         reasonOutputSwitchedOff2 : Int;   // 0=output current>limit and output current<1,5xlimit for more than 5sec; 1=current output>1,5xlimit; 2=total overload; 3=Uin<19,4V and output current>limit; 4=Uin<15V; 5=Uin>30V; 6=device overtemperature; 8 to 14=Reserve; 15=default (no automatically switched off)
         reasonOutputSwitchedOff3 : Int;   // 0=output current>limit and output current<1,5xlimit for more than 5sec; 1=current output>1,5xlimit; 2=total overload; 3=Uin<19,4V and output current>limit; 4=Uin<15V; 5=Uin>30V; 6=device overtemperature; 8 to 14=Reserve; 15=default (no automatically switched off)
         reasonOutputSwitchedOff4 : Int;   // 0=output current>limit and output current<1,5xlimit for more than 5sec; 1=current output>1,5xlimit; 2=total overload; 3=Uin<19,4V and output current>limit; 4=Uin<15V; 5=Uin>30V; 6=device overtemperature; 8 to 14=Reserve; 15=default (no automatically switched off)
         reasonOutputSwitchedOff5 : Int;   // 0=output current>limit and output current<1,5xlimit for more than 5sec; 1=current output>1,5xlimit; 2=total overload; 3=Uin<19,4V and output current>limit; 4=Uin<15V; 5=Uin>30V; 6=device overtemperature; 8 to 14=Reserve; 15=default (no automatically switched off)
         reasonOutputSwitchedOff6 : Int;   // 0=output current>limit and output current<1,5xlimit for more than 5sec; 1=current output>1,5xlimit; 2=total overload; 3=Uin<19,4V and output current>limit; 4=Uin<15V; 5=Uin>30V; 6=device overtemperature; 8 to 14=Reserve; 15=default (no automatically switched off)
         reasonOutputSwitchedOff7 : Int;   // 0=output current>limit and output current<1,5xlimit for more than 5sec; 1=current output>1,5xlimit; 2=total overload; 3=Uin<19,4V and output current>limit; 4=Uin<15V; 5=Uin>30V; 6=device overtemperature; 8 to 14=Reserve; 15=default (no automatically switched off)
         reasonOutputSwitchedOff8 : Int;   // 0=output current>limit and output current<1,5xlimit for more than 5sec; 1=current output>1,5xlimit; 2=total overload; 3=Uin<19,4V and output current>limit; 4=Uin<15V; 5=Uin>30V; 6=device overtemperature; 8 to 14=Reserve; 15=default (no automatically switched off)
         nominalOutputCurrent : Int;   // nominal output current
         outputNumber : Int;   // number of outputs (4 or 8)
         productState : Int;   // product state
         firmwareVersion : Int;   // frimware version
         startup : Int;   // 0=load dependent startup; 1=startup time tag 25ms; 2=startup time tag 200ms; 3=startup time tag 500ms
         setReset : Bool;
         stateReset : Bool;
         stateNoCommunication : Bool;
         articleNumber : String;   // article number
         serialNumber : String;   // serial number
      END_STRUCT;
      statIndexResetBitArray : Int;
      statInit : Bool;
      statArticleNumber : Array[1..18] of Char;
      statArticleNumberOld : Array[1..18] of Char;
      statSerialNumber : Array[1..13] of Char;
      statSerialNumberOld : Array[1..13] of Char;
      statVarianten11String : String[2];
      statInnovationenString : String[2];
      statArticleNumberChanged : Bool;
      statErrorFrameContent : Bool;
      statErrorFrameID : Bool;
      statErrorFrameLength : Bool;
      statErrorDevice : Bool;
      statIndexArticleNumber : Int := 1;
      statIndexSerialNumber : Int := 1;
      statNewArticleNumberDetected : Bool;
      statNewSerialNumberDetected : Bool;
      instTimerReset : TON_TIME;
      statCntReason : Int;
      statCntCurrentLimit : Int;
   END_VAR
   VAR_TEMP
      tempLatchTime : Time;
      tempRetval : Word;
      tempRetvalSysTime : Int;
      tempRetvalSysPosEdge : Int;
      tempRetvalSysNegEdge : Int;
   END_VAR
   VAR CONSTANT
      CONST_POS_EDGE : Int := 15;
      CONST_NEG_EDGE : Int := 16;
      STATE_IDLE : Int := 1;
      STATE_EVALUATION : Int := 2;
      STATE_ERROR : Int := 3;
      CONST_DWORD_0 : DWord := 16#0000_0000;
      CONST_WORD_0 : Word := 16#0000;
      CONST_BYTE_0 : Byte := 16#00;
      CONST_INT_0 : Int := 0;
      CONST_INT_1 : Int := 1;
      CONST_TIME_0 : Time := T#0MS;
      CONST_TIME_WAIT : Time := T#65MS;
      CONST_SYS_TIMER : Time := T#4S;
      CONST_WATCHDOG_TIMER : Time := T#9S;
      CONST_INIT_TIMER : Time := T#4S;
      CONST_RESET_TIMER : Time := T#50ms;
      CONST_START_IMPULSE_MIN : Time := T#126MS;
      CONST_START_IMPULSE_MAX : Time := T#175MS;
      CONST_IMPULSE_MIN : Time := T#25MS;
      CONST_IMPULSE_MAX : Time := T#125MS;
      CONST_PAUSE_MAX : Time := T#125MS;
      CONST_PAUSE_MIN : Time := T#25MS;
      CONST_START_CNT_INDEX0 : Int := 0;
      CONST_START_CNT_INDEX1 : Int := 1;
      CONST_END_CNT_INDEX63 : Int := 63;
      CONST_END_CNT_INDEX31 : Int := 31;
      CONST_END_CNT_INDEX18 : Int := 18;
      CONST_END_CNT_INDEX13 : Int := 13;
      CONST_FRAME_MAX : Time := T#3S_625MS;
      CONST_FRAME_MIN : Time := T#3S_275MS;
      CONST_CNT_BITS_MAX : Int := 32;
      CONST_CNT_PAUSE_MAX : Int := 33;
      CONST_TIME_CYCLE_MAX : Time := T#12MS;
      CONST_ERR_ARTICLE_NUMBER : Word := 16#8007;
      CONST_ERR_FRAME_ID : Word := 16#8006;
      CONST_ERR_DEVICE : Word := 16#8005;
      CONST_ERR_FRAMELENGTH : Word := 16#8004;
      CONST_ERR_FRAMECONTENT : Word := 16#8003;
      CONST_ERR_CYCLE_TIME : Word := 16#8002;
      CONST_ERR_WATCHDOG : Word := 16#8001;
      CONST_CONVERT_CURRENT : Int := 10;
      CONST_NOMINAL_VALUE_DETECT0 : Byte := 16#00;
      CONST_NOMINAL_VALUE_DETECT1 : Byte := 16#01;
      CONST_NOMINAL_VALUE_DETECT2 : Byte := 16#02;
      CONST_NOMINAL_CURRENT3 : Int := 3;
      CONST_NOMINAL_CURRENT5 : Int := 5;
      CONST_NOMINAL_CURRENT10 : Int := 10;
      CONST_NOMINAL_VOLTAGE : Int := 24;
      CONST_YEAR_2019 : Int := 2019;
      CONST_YEAR_2020 : Int := 2020;
      CONST_YEAR_2021 : Int := 2021;
      CONST_YEAR_2022 : Int := 2022;
      CONST_YEAR_2023 : Int := 2023;
      CONST_YEAR_2024 : Int := 2024;
      CONST_YEAR_2025 : Int := 2025;
      CONST_YEAR_2026 : Int := 2026;
      CONST_YEAR_2027 : Int := 2027;
      CONST_YEAR_2028 : Int := 2028;
      CONST_YEAR_2029 : Int := 2029;
      CONST_YEAR_2030 : Int := 2030;
      CONST_YEAR_2031 : Int := 2031;
      CONST_YEAR_2032 : Int := 2032;
      CONST_YEAR_2033 : Int := 2033;
      CONST_YEAR_2034 : Int := 2034;
      CONST_FRAME_ID0 : Int := 0;
      CONST_FRAME_ID1 : Int := 1;
      CONST_FRAME_ID2 : Int := 2;
      CONST_FRAME_ID3 : Int := 3;
      CONST_DEVICE_SEL1200 : Int := 1;
      CONST_DEVICE_SEL1400 : Int := 2;
      CONST_JANUARY : Int := 1;
      CONST_FEBRUARY : Int := 2;
      CONST_MARCH : Int := 3;
      CONST_APRIL : Int := 4;
      CONST_MAY : Int := 5;
      CONST_JUNE : Int := 6;
      CONST_JULY : Int := 7;
      CONST_AUGUST : Int := 8;
      CONST_SEPTEMBER : Int := 9;
      CONST_OCTOBER : Int := 10;
      CONST_NOVEMBER : Int := 11;
      CONST_DECEMBER : Int := 12;
      CONST_ONE_CHANNEL : Int := 0;
      CONST_TWO_CHANNEL : Int := 1;
      CONST_FOUR_CHANNEL : Int := 2;
      CONST_EIGHT_CHANNEL : Int := 3;
      CONST_NO_DESCRIPTION : Int := 4;
      CONST_GLITCH_MAX : Int := 32000;
      CONST_MEASUREMENT_CURRENT : Int := 0;
      CONST_MEASUREMENT_CURRENT_LIMIT : Int := 2;
      CONST_OUTPUT_NUMBER_4 : Int := 4;
      CONST_OUTPUT_NUMBER_8 : Int := 8;
      CONST_POWER_0 : Int := 0;
      CONST_POWER_20 : Int := 20;
      CONST_POWER_50 : Int := 50;
      CONST_POWER_100 : Int := 100;
      CONST_POWER_150 : Int := 150;
      CONST_POWER_250 : Int := 250;
      CONST_POWER_400 : Int := 400;
      CONST_POWER_600 : Int := 600;
      CONST_POWER_1000 : Int := 100;
      CONST_REASON_DEFAULT : Int := 0;
      CONST_STATE_OUT_AUTO_SWITCHED_OFF : Int := 0;
      CONST_STATE_OUT_RESET_POSSIBLE : Int := 1;
      CONST_DEVICE_NAME_DEFAULT : String := 'SEL1200';
      CONST_ARTICLE_NUMBER_DEFAULT : String := '6EP4437-7FB00-0CX0';
      CONST_SERIAL_NUMBER_DEFAULT : String := 'Q6/L1';
      CONST_STATE_OUT_DEFAULT : Int := 0;
      CONST_CURRENT_OUT_DEFAULT : Int := 0;
      CONST_REASON_SWITCHED_OFF_DEFAULT : Int := 0;
      CONST_FW_PRODUCT_STATE_DEFAULT : Int := 1;
      CONST_STARTUP_DEFAULT : Int := 0;
   END_VAR
BEGIN

REGION Network 1 (SCL)
   //=============================================================================
   //SIEMENES AG
   //(c)Copyright 2019 All Rights Reserved
   //-----------------------------------------------------------------------------
   //Library:       LPSU6200_V15.0-0_V1-0-0
   //Tested with:   (S7-1500)
   //Engineering:    TIA Portal V15
   //Restrictions:   call in cyclic interrupt OB with max. 10ms
   //Requirements:
   //Functionality: evaluates the signal of diagnostic interface of SITOP PSU6200 
   //               ....
   //
   //-----------------------------------------------------------------------------
   //Change log table:
   //Version  Date       Expert in charge Changes applied
   //01.00.00 17.01.2019 (DF CS SD CSS KMT KD) First released version
   //=============================================================================


   // Calculate cycle time
   #tempRetvalSysTime := RD_SYS_T(#statTimeSave.sysTime);

   IF #statTimeSave.sysTime > #statTimeSave.sysTimeOld
   THEN
       //Calculate cycle time
       #statTimeSave.deltaSysTime := T_DIFF(IN1 := #statTimeSave.sysTime,
                                            IN2 := #statTimeSave.sysTimeOld);
       #statStartTimerSys := false;
   ELSE
       #statStartTimerSys := true;
       #statTimeSave.sysTimeOld := #statTimeSave.sysTime;
       RETURN;
   END_IF;

   //check cycle time

   IF (#statTimeSave.deltaSysTime >= #CONST_TIME_CYCLE_MAX)
   THEN
       #statCycleTimeNotOk := true;
       #statStartTimerSys := true;
   ELSE
       #statCycleTimeNotOk := false;
       #statStartTimerSys := false;
   END_IF;


   //pos edge detection

   IF #impulse = TRUE
       AND #statImpulseOld = FALSE
   THEN
       #tempRetvalSysPosEdge := RD_SYS_T(#statTimeSave.posEdge);
       #statPosEdgeDetected := true;
       #statPosEdgeDetectedTrigger := true;
       #statEdgeCtrl := #CONST_POS_EDGE;
       #statStartWatchDogTimerPos := true;
       #statStartWatchDogTimerNeg := false;
       #HMI.stateNoCommunication := false;

       IF #statBusy = FALSE
       THEN
           #statInit := false;
           #statBusy := true;
           #statDone := false;
           #statError := false;
           #statStatus := #CONST_WORD_0;
       END_IF;

       IF #statCycleTimeNotOk = FALSE
       THEN
           #statStateIndex := #STATE_EVALUATION;
       END_IF;

   END_IF;

   //neg edge detection

   IF #impulse = false
       AND #statImpulseOld = true
   THEN
       #tempRetvalSysNegEdge := RD_SYS_T(#statTimeSave.negEdge);
       #statNegEdgeDetected := true;
       #statNegEdgeDetectedTrigger := true;
       #statEdgeCtrl := #CONST_NEG_EDGE;
       #statStartWatchDogTimerNeg := true;
       #statStartWatchDogTimerPos := false;

       IF #statCycleTimeNotOk = FALSE
       THEN
           #statStateIndex := #STATE_EVALUATION;
       END_IF;

   END_IF;

   IF #statPosEdgeDetected = FALSE
       AND #statNegEdgeDetected = FALSE
   THEN
       #statStartWatchDogTimerPos := true;
       #statStartWatchDogTimerNeg := true;
   END_IF;


   CASE #statStateIndex OF
       #STATE_IDLE:  // State IDLE

           #statError := false;
           #statErrorInt := false;
           #statDone := false;
           #statBusy := false;
           #statStatus := #CONST_WORD_0;
           #statFrame := #CONST_DWORD_0;
           #statInit := false;
           #error := false;
           #done := false;
           #busy := false;
           #status := #CONST_WORD_0;
           #frame := #CONST_DWORD_0;

           #statNoEvaluation := false;
           #statFrameEvaluationStopp := false;
           #statStartTimerWait := false;
           #statCycleTimeNotOk := false;
           #statPosEdgeDetected := false;
           #statNegEdgeDetected := false;
           #HMI.stateNoCommunication := false;

           FOR #statIndexResetBitArray := #CONST_START_CNT_INDEX0 TO #CONST_END_CNT_INDEX31 DO
               // Statement section FOR
               #statArrayBits[#statIndexResetBitArray] := false;
           END_FOR;


       #STATE_EVALUATION:

           IF #statPosEdgeDetected = TRUE
               AND #statNegEdgeDetected = true
           THEN


               // Delta Time calculation

               IF #statEdgeCtrl = #CONST_POS_EDGE
               THEN
                   #statPauseDetected := true;

                   // time of pause
                   #statTimeSave.deltaTimePause := T_DIFF(IN1 := #statTimeSave.posEdge,
                                                          IN2 := #statTimeSave.negEdge);

                   //check time of pause
                   IF #statTimeSave.deltaTimePause < #CONST_TIME_0
                   THEN
                       #statErrorFrameContent := TRUE;
                   ELSIF (#statTimeSave.deltaTimePause < #CONST_PAUSE_MIN)
                       OR (#statTimeSave.deltaTimePause > #CONST_PAUSE_MAX)
                   THEN
                       #statErrorFrameContent := TRUE;
                   END_IF;

                   #statNegEdgeDetected := false;
               END_IF;

               IF #statEdgeCtrl = #CONST_NEG_EDGE
               THEN
                   #statImpulseDetected := true;

                   // time of impulse
                   #statTimeSave.deltaTimeImpulse := T_DIFF(IN1 := #statTimeSave.negEdge,
                                                            IN2 := #statTimeSave.posEdge);

                   //check time of impulse

                   IF #statTimeSave.deltaTimeImpulse < #CONST_TIME_0
                   THEN
                       #statErrorFrameContent := TRUE;

                   ELSIF (#statTimeSave.deltaTimeImpulse < #CONST_IMPULSE_MIN)
                       OR (#statTimeSave.deltaTimeImpulse > #CONST_START_IMPULSE_MAX)
                   THEN
                       #statErrorFrameContent := TRUE;
                   END_IF;

                   #statPosEdgeDetected := false;
               END_IF;

           END_IF;

           //Startbit detection
           IF (#statTimeSave.deltaTimeImpulse >= #CONST_START_IMPULSE_MIN)
               AND (#statTimeSave.deltaTimeImpulse <= #CONST_START_IMPULSE_MAX)
               AND (#statImpulseDetected = true)
           THEN
               #statImpulseDetected := false;
               #statIndexImpulse := #CONST_INT_1;
               #statIndexPause := #CONST_INT_0;
               #statFrameEvaluationStopp := false;
               #statCntBits := #CONST_INT_0;
               #statCntImpulse := #CONST_INT_0;
               #statCntPause := #CONST_INT_0;
               #statTimeSave.timeIpulse := #CONST_TIME_0;
               #statTimeSave.timePause := #CONST_TIME_0;
               #statIndexAddTime := #CONST_INT_0;

               //check frame length
               FOR #statIndexAddTime := #CONST_START_CNT_INDEX0 TO #CONST_END_CNT_INDEX63 BY 1 DO
                   #statTimeSave.timeIpulse := #statTimeSave.timeIpulse + #statArrayImpulse[#statIndexAddTime];
                   #statTimeSave.timePause := #statTimeSave.timePause + #statArrayPause[#statIndexAddTime];
               END_FOR;

               #statTimeSave.timeFrame := #statTimeSave.timeIpulse + #statTimeSave.timePause;

               IF #statTimeSave.timeFrame >= #CONST_FRAME_MIN
                   AND #statTimeSave.timeFrame <= #CONST_FRAME_MAX
               THEN
                   //CollectData

                   #statDone := true;
                   #statBusy := false;
                   #statInit := true;

                   #statFrame.%X0 := #statArrayBits[0];
                   #statFrame.%X1 := #statArrayBits[1];
                   #statFrame.%X2 := #statArrayBits[2];
                   #statFrame.%X3 := #statArrayBits[3];
                   #statFrame.%X4 := #statArrayBits[4];
                   #statFrame.%X5 := #statArrayBits[5];
                   #statFrame.%X6 := #statArrayBits[6];
                   #statFrame.%X7 := #statArrayBits[7];
                   #statFrame.%X8 := #statArrayBits[8];
                   #statFrame.%X9 := #statArrayBits[9];
                   #statFrame.%X10 := #statArrayBits[10];
                   #statFrame.%X11 := #statArrayBits[11];
                   #statFrame.%X12 := #statArrayBits[12];
                   #statFrame.%X13 := #statArrayBits[13];
                   #statFrame.%X14 := #statArrayBits[14];
                   #statFrame.%X15 := #statArrayBits[15];
                   #statFrame.%X16 := #statArrayBits[16];
                   #statFrame.%X17 := #statArrayBits[17];
                   #statFrame.%X18 := #statArrayBits[18];
                   #statFrame.%X19 := #statArrayBits[19];
                   #statFrame.%X20 := #statArrayBits[20];
                   #statFrame.%X21 := #statArrayBits[21];
                   #statFrame.%X22 := #statArrayBits[22];
                   #statFrame.%X23 := #statArrayBits[23];
                   #statFrame.%X24 := #statArrayBits[24];
                   #statFrame.%X25 := #statArrayBits[25];
                   #statFrame.%X26 := #statArrayBits[26];
                   #statFrame.%X27 := #statArrayBits[27];
                   #statFrame.%X28 := #statArrayBits[28];
                   #statFrame.%X29 := #statArrayBits[29];
                   #statFrame.%X30 := #statArrayBits[30];
                   #statFrame.%X31 := #statArrayBits[31];

                   #frame := #statFrame;

                   IF #statFrame <> #statFrameOld
                   THEN


                       #statDeviceName.%X2 := #statFrame.%X0;
                       #statDeviceName.%X1 := #statFrame.%X1;
                       #statDeviceName.%X0 := #statFrame.%X2;

                       //device detection 
                       //SEL1200 or SEL1400
                       IF (BYTE_TO_INT(#statDeviceName) = #CONST_DEVICE_SEL1200)
                           OR (BYTE_TO_INT(#statDeviceName) = #CONST_DEVICE_SEL1400)
                       THEN
                           IF BYTE_TO_INT(#statDeviceName) = #CONST_DEVICE_SEL1200
                           THEN
                               #statHMI.deviceName := 'SEL1200';
                               #statArticleNumber[10] := 'F'; // constant value pos 9
                           ELSIF BYTE_TO_INT(#statDeviceName) = #CONST_DEVICE_SEL1400
                           THEN
                               #statHMI.deviceName := 'SEL1400';
                               #statArticleNumber[10] := 'E'; // constant value pos 9
                           END_IF;

                           #statArticleNumber[1] := '6';  // constant value pos 1
                           #statArticleNumber[2] := 'E';  // constant value pos 2
                           #statArticleNumber[3] := 'P';  // constant value pos 3
                           #statArticleNumber[4] := '4';  // device SEL1200 or SEL1400 (sectivity module) pos 4
                           #statArticleNumber[5] := '4';  // family (diagnostic module) pos 5
                           #statArticleNumber[6] := '3';  // output voltage <=24V DC, constant value pos 6 
                           #statArticleNumber[8] := '-';  // constant value
                           #statArticleNumber[9] := '7';  // constant value pos 8
                           #statArticleNumber[14] := '-';  // constant value
                           #statArticleNumber[15] := '3';  // constant value pos 13 (interface: messages in Morse code)
                           #statArticleNumber[17] := 'X';  // constant value pos 15
                           #statArticleNumber[18] := '0';  // constant value pos 16

                           //FrameId detection
                           #statFrameID.%X1 := #statFrame.%X4;
                           #statFrameID.%X0 := #statFrame.%X5;

                           //state information channel 1 to 8

                           IF BYTE_TO_INT(#statFrameID) = #CONST_FRAME_ID0
                           THEN
                               #statGetFrame.frame0 := true;

                               // state input voltage 
                               #statStateInputVoltage := #statFrame.%X6; //0= input voltage to low or high; 1: input voltage ok

                               //state channel 1
                               //0: channel is switched off automatically, no reset possible
                               //1: channel is switched off automatically, reset possible
                               //2: channel is switched off manually
                               //3: channel is sitched on
                               //4: channel is defect
                               //5: device overtemperature, channel is switched off
                               //6: overload, in sum the current of all channels to high
                               //7: current of channel is higher than nominal current
                               #statStateOutput1.%X2 := #statFrame.%X7;
                               #statStateOutput1.%X1 := #statFrame.%X8;
                               #statStateOutput1.%X0 := #statFrame.%X9;
                               #statHMI.stateOutput1 := BYTE_TO_INT(#statStateOutput1);

                               IF (#statHMI.stateOutput1 <> #CONST_STATE_OUT_AUTO_SWITCHED_OFF)
                                   AND (#statHMI.stateOutput1 <> #CONST_STATE_OUT_RESET_POSSIBLE)
                               THEN
                                   #statHMI.reasonOutputSwitchedOff1 := #CONST_REASON_DEFAULT;
                               END_IF;

                               //state channel 2
                               #statStateOutput2.%X2 := #statFrame.%X10;
                               #statStateOutput2.%X1 := #statFrame.%X11;
                               #statStateOutput2.%X0 := #statFrame.%X12;
                               #statHMI.stateOutput2 := BYTE_TO_INT(#statStateOutput2);

                               IF (#statHMI.stateOutput2 <> #CONST_STATE_OUT_AUTO_SWITCHED_OFF)
                                   AND (#statHMI.stateOutput2 <> #CONST_STATE_OUT_RESET_POSSIBLE)
                               THEN
                                   #statHMI.reasonOutputSwitchedOff2 := #CONST_REASON_DEFAULT;
                               END_IF;

                               //state channel 3
                               #statStateOutput3.%X2 := #statFrame.%X13;
                               #statStateOutput3.%X1 := #statFrame.%X14;
                               #statStateOutput3.%X0 := #statFrame.%X15;
                               #statHMI.stateOutput3 := BYTE_TO_INT(#statStateOutput3);

                               IF (#statHMI.stateOutput3 <> #CONST_STATE_OUT_AUTO_SWITCHED_OFF)
                                   AND (#statHMI.stateOutput3 <> #CONST_STATE_OUT_RESET_POSSIBLE)
                               THEN
                                   #statHMI.reasonOutputSwitchedOff3 := #CONST_REASON_DEFAULT;
                               END_IF;

                               //state channel 4
                               #statStateOutput4.%X2 := #statFrame.%X16;
                               #statStateOutput4.%X1 := #statFrame.%X17;
                               #statStateOutput4.%X0 := #statFrame.%X18;
                               #statHMI.stateOutput4 := BYTE_TO_INT(#statStateOutput4);

                               IF (#statHMI.stateOutput4 <> #CONST_STATE_OUT_AUTO_SWITCHED_OFF)
                                   AND (#statHMI.stateOutput4 <> #CONST_STATE_OUT_RESET_POSSIBLE)
                               THEN
                                   #statHMI.reasonOutputSwitchedOff4 := #CONST_REASON_DEFAULT;
                               END_IF;

                               //state channel 5
                               #statStateOutput5.%X2 := #statFrame.%X19;
                               #statStateOutput5.%X1 := #statFrame.%X20;
                               #statStateOutput5.%X0 := #statFrame.%X21;
                               #statHMI.stateOutput5 := BYTE_TO_INT(#statStateOutput5);

                               IF (#statHMI.stateOutput5 <> #CONST_STATE_OUT_AUTO_SWITCHED_OFF)
                                   AND (#statHMI.stateOutput5 <> #CONST_STATE_OUT_RESET_POSSIBLE)
                               THEN
                                   #statHMI.reasonOutputSwitchedOff5 := #CONST_REASON_DEFAULT;
                               END_IF;

                               //state channel 6
                               #statStateOutput6.%X2 := #statFrame.%X22;
                               #statStateOutput6.%X1 := #statFrame.%X23;
                               #statStateOutput6.%X0 := #statFrame.%X24;
                               #statHMI.stateOutput6 := BYTE_TO_INT(#statStateOutput6);

                               IF (#statHMI.stateOutput6 <> #CONST_STATE_OUT_AUTO_SWITCHED_OFF)
                                   AND (#statHMI.stateOutput6 <> #CONST_STATE_OUT_RESET_POSSIBLE)
                               THEN
                                   #statHMI.reasonOutputSwitchedOff6 := #CONST_REASON_DEFAULT;
                               END_IF;

                               //state channel 7
                               #statStateOutput7.%X2 := #statFrame.%X25;
                               #statStateOutput7.%X1 := #statFrame.%X26;
                               #statStateOutput7.%X0 := #statFrame.%X27;
                               #statHMI.stateOutput7 := BYTE_TO_INT(#statStateOutput7);

                               IF (#statHMI.stateOutput7 <> #CONST_STATE_OUT_AUTO_SWITCHED_OFF)
                                   AND (#statHMI.stateOutput7 <> #CONST_STATE_OUT_RESET_POSSIBLE)
                               THEN
                                   #statHMI.reasonOutputSwitchedOff7 := #CONST_REASON_DEFAULT;
                               END_IF;

                               //state channel 8
                               #statStateOutput8.%X2 := #statFrame.%X28;
                               #statStateOutput8.%X1 := #statFrame.%X29;
                               #statStateOutput8.%X0 := #statFrame.%X30;
                               #statHMI.stateOutput8 := BYTE_TO_INT(#statStateOutput8);

                               IF (#statHMI.stateOutput8 <> #CONST_STATE_OUT_AUTO_SWITCHED_OFF)
                                   AND (#statHMI.stateOutput8 <> #CONST_STATE_OUT_RESET_POSSIBLE)
                               THEN
                                   #statHMI.reasonOutputSwitchedOff8 := #CONST_REASON_DEFAULT;
                               END_IF;

                               IF #statHMI.stateOutput1 = #CONST_STATE_OUT_RESET_POSSIBLE
                                   OR #statHMI.stateOutput2 = #CONST_STATE_OUT_RESET_POSSIBLE
                                   OR #statHMI.stateOutput3 = #CONST_STATE_OUT_RESET_POSSIBLE
                                   OR #statHMI.stateOutput4 = #CONST_STATE_OUT_RESET_POSSIBLE
                                   OR #statHMI.stateOutput5 = #CONST_STATE_OUT_RESET_POSSIBLE
                                   OR #statHMI.stateOutput6 = #CONST_STATE_OUT_RESET_POSSIBLE
                                   OR #statHMI.stateOutput7 = #CONST_STATE_OUT_RESET_POSSIBLE
                                   OR #statHMI.stateOutput8 = #CONST_STATE_OUT_RESET_POSSIBLE
                               THEN
                                   #statHMI.stateReset := true;
                               ELSE
                                   #statHMI.stateReset := false;
                               END_IF;

                               // device data
                           ELSIF
                               BYTE_TO_INT(#statFrameID) = #CONST_FRAME_ID1
                           THEN
                               #statGetFrame.frame1 := true;

                               //Construction Month
                               #statConstructionMonthByte.%X3 := #statFrame.%X6;
                               #statConstructionMonthByte.%X2 := #statFrame.%X7;
                               #statConstructionMonthByte.%X1 := #statFrame.%X8;
                               #statConstructionMonthByte.%X0 := #statFrame.%X9;
                               #statConstructionMonth := BYTE_TO_INT(#statConstructionMonthByte);

                               IF #statConstructionMonth = #CONST_JANUARY //January
                               THEN
                                   #statConstructionMonthChar := '1';
                               ELSIF #statConstructionMonth = #CONST_FEBRUARY //February
                               THEN
                                   #statConstructionMonthChar := '2';
                               ELSIF #statConstructionMonth = #CONST_MARCH //March
                               THEN
                                   #statConstructionMonthChar := '3';
                               ELSIF #statConstructionMonth = #CONST_APRIL //April
                               THEN
                                   #statConstructionMonthChar := '4';
                               ELSIF #statConstructionMonth = #CONST_MAY // May
                               THEN
                                   #statConstructionMonthChar := '5';
                               ELSIF #statConstructionMonth = #CONST_JUNE //June
                               THEN
                                   #statConstructionMonthChar := '6';
                               ELSIF #statConstructionMonth = #CONST_JULY //July
                               THEN
                                   #statConstructionMonthChar := '7';
                               ELSIF #statConstructionMonth = #CONST_AUGUST //August
                               THEN
                                   #statConstructionMonthChar := '8';
                               ELSIF #statConstructionMonth = #CONST_SEPTEMBER //September
                               THEN
                                   #statConstructionMonthChar := '9';
                               ELSIF #statConstructionMonth = #CONST_OCTOBER //October
                               THEN
                                   #statConstructionMonthChar := '0';
                               ELSIF #statConstructionMonth = #CONST_NOVEMBER // November
                               THEN
                                   #statConstructionMonthChar := 'N';
                               ELSIF #statConstructionMonth = #CONST_DECEMBER //December
                               THEN
                                   #statConstructionMonthChar := 'D';
                               ELSE
                                   #statConstructionMonthChar := '1';

                               END_IF;

                               //Software Version
                               #statFirmwareVersion.%X2 := #statFrame.%X10;
                               #statFirmwareVersion.%X1 := #statFrame.%X11;
                               #statFirmwareVersion.%X0 := #statFrame.%X12;
                               #statHMI.firmwareVersion := BYTE_TO_INT(#statFirmwareVersion);

                               //Varianten for article number pos 11
                               #statVarianten11.%X2 := #statFrame.%X13;
                               #statVarianten11.%X1 := #statFrame.%X14;
                               #statVarianten11.%X0 := #statFrame.%X15;

                               #tempRetval := HTA(IN := #statVarianten11, N := 1, OUT => #statVarianten11String);
                               #statVarianten11String := DELETE(IN := #statVarianten11String, L := 1, P := 1);
                               #statArticleNumber[12] := #statVarianten11String;

                               //Inovationen for article number pos 12
                               #statInnovationen.%X2 := #statFrame.%X16;
                               #statInnovationen.%X1 := #statFrame.%X17;
                               #statInnovationen.%X0 := #statFrame.%X18;

                               #tempRetval := HTA(IN := #statInnovationen, N := 1, OUT => #statInnovationenString);
                               #statInnovationenString := DELETE(IN := #statInnovationenString, L := 1, P := 1);
                               #statArticleNumber[13] := #statInnovationenString;

                               //number of channels for article number pos 14
                               #statChannelNumber.%X2 := #statFrame.%X19;
                               #statChannelNumber.%X1 := #statFrame.%X20;
                               #statChannelNumber.%X0 := #statFrame.%X21;

                               // for article number pos. 14
                               IF BYTE_TO_INT(#statChannelNumber) = #CONST_ONE_CHANNEL
                               THEN
                                   #statArticleNumber[16] := 'A'; //one channel
                               ELSIF
                                   BYTE_TO_INT(#statChannelNumber) = #CONST_TWO_CHANNEL
                               THEN
                                   #statArticleNumber[16] := 'B'; // two channels
                               ELSIF BYTE_TO_INT(#statChannelNumber) = #CONST_FOUR_CHANNEL
                               THEN
                                   #statArticleNumber[16] := 'C'; // four channels
                               ELSIF BYTE_TO_INT(#statChannelNumber) = #CONST_EIGHT_CHANNEL
                               THEN
                                   #statArticleNumber[16] := 'D'; // eight channels
                               ELSIF BYTE_TO_INT(#statChannelNumber) = #CONST_NO_DESCRIPTION
                               THEN
                                   #statArticleNumber[16] := 'X'; //no description
                               ELSE
                                   // default value
                                   #statArticleNumber[16] := 'A';
                               END_IF;

                               //Construction Year
                               #statConstructionYearByte.%X3 := #statFrame.%X22;
                               #statConstructionYearByte.%X2 := #statFrame.%X23;
                               #statConstructionYearByte.%X1 := #statFrame.%X24;
                               #statConstructionYearByte.%X0 := #statFrame.%X25;

                               #statConstructionYear := BYTE_TO_INT(#statConstructionYearByte) + #CONST_YEAR_2019;

                               IF #statConstructionYear = #CONST_YEAR_2019
                               THEN
                                   #statConstructionYearChar := 'L';
                               ELSIF #statConstructionYear = #CONST_YEAR_2020
                               THEN
                                   #statConstructionYearChar := 'M';
                               ELSIF #statConstructionYear = #CONST_YEAR_2021
                               THEN
                                   #statConstructionYearChar := 'N';
                               ELSIF #statConstructionYear = #CONST_YEAR_2022
                               THEN
                                   #statConstructionYearChar := 'P';
                               ELSIF #statConstructionYear = #CONST_YEAR_2023
                               THEN
                                   #statConstructionYearChar := 'R';
                               ELSIF #statConstructionYear = #CONST_YEAR_2024
                               THEN
                                   #statConstructionYearChar := 'S';
                               ELSIF #statConstructionYear = #CONST_YEAR_2025
                               THEN
                                   #statConstructionYearChar := 'T';
                               ELSIF #statConstructionYear = #CONST_YEAR_2026
                               THEN
                                   #statConstructionYearChar := 'U';
                               ELSIF #statConstructionYear = #CONST_YEAR_2027
                               THEN
                                   #statConstructionYearChar := 'V';
                               ELSIF #statConstructionYear = #CONST_YEAR_2028
                               THEN
                                   #statConstructionYearChar := 'W';
                               ELSIF #statConstructionYear = #CONST_YEAR_2029
                               THEN
                                   #statConstructionYearChar := 'X';
                               ELSIF #statConstructionYear = #CONST_YEAR_2030
                               THEN
                                   #statConstructionYearChar := 'A';
                               ELSIF #statConstructionYear = #CONST_YEAR_2031
                               THEN
                                   #statConstructionYearChar := 'B';
                               ELSIF #statConstructionYear = #CONST_YEAR_2032
                               THEN
                                   #statConstructionYearChar := 'C';
                               ELSIF #statConstructionYear = #CONST_YEAR_2033
                               THEN
                                   #statConstructionYearChar := 'D';
                               ELSIF #statConstructionYear = #CONST_YEAR_2034
                               THEN
                                   #statConstructionYearChar := 'E';
                               ELSE
                                   #statConstructionYearChar := 'L';
                               END_IF;

                               //Product Version
                               #statProductState.%X2 := #statFrame.%X26;
                               #statProductState.%X1 := #statFrame.%X27;
                               #statProductState.%X0 := #statFrame.%X28;

                               #statHMI.productState := BYTE_TO_INT(#statProductState);

                               //normal or lacquered
                               #statLacquered := #statFrame.%X29;

                               IF #statLacquered = TRUE
                               THEN
                                   #statArticleNumber[11] := 'C';  //article number pos 10
                               ELSE
                                   #statArticleNumber[11] := 'B'; //article number pos 10
                               END_IF;

                               //fabrication place
                               #statFabricationPlace := #statFrame.%X30;


                           ELSIF BYTE_TO_INT(#statFrameID) = #CONST_FRAME_ID2
                           THEN

                               #statGetFrame.frame2 := true;

                               #statMeasurementsChannels.%X1 := #statFrame.%X6;
                               #statMeasurementsChannels.%X0 := #statFrame.%X7;


                               IF BYTE_TO_INT(#statMeasurementsChannels) = #CONST_MEASUREMENT_CURRENT
                               THEN
                                   //measurement output current (channel 1 to 4)
                                   #statGetFrame.frame21 := true;

                                   //current output 1 (0% to 150% of nominal value)
                                   #statOutputCurrent1.%X3 := #statFrame.%X8;
                                   #statOutputCurrent1.%X2 := #statFrame.%X9;
                                   #statOutputCurrent1.%X1 := #statFrame.%X10;
                                   #statOutputCurrent1.%X0 := #statFrame.%X11;

                                   //current output 2 (0% to 150% of nominal value)
                                   #statOutputCurrent2.%X3 := #statFrame.%X12;
                                   #statOutputCurrent2.%X2 := #statFrame.%X13;
                                   #statOutputCurrent2.%X1 := #statFrame.%X14;
                                   #statOutputCurrent2.%X0 := #statFrame.%X15;

                                   //current output 3 (0% to 150% of nominal value)
                                   #statOutputCurrent3.%X3 := #statFrame.%X16;
                                   #statOutputCurrent3.%X2 := #statFrame.%X17;
                                   #statOutputCurrent3.%X1 := #statFrame.%X18;
                                   #statOutputCurrent3.%X0 := #statFrame.%X19;

                                   //current output 4 (0% to 150% of nominal value)
                                   #statOutputCurrent4.%X3 := #statFrame.%X20;
                                   #statOutputCurrent4.%X2 := #statFrame.%X21;
                                   #statOutputCurrent4.%X1 := #statFrame.%X22;
                                   #statOutputCurrent4.%X0 := #statFrame.%X23;

                               ELSIF BYTE_TO_INT(#statMeasurementsChannels) = #CONST_MEASUREMENT_CURRENT_LIMIT
                               THEN
                                   // output current limit on potentiometer (channel 1 to 4)
                                   #statGetFrame.frame22 := true;

                                   //current limit of output 1 (0% to 100% of nominal value)
                                   #statOutputCurrentLimit1.%X3 := #statFrame.%X8;
                                   #statOutputCurrentLimit1.%X2 := #statFrame.%X9;
                                   #statOutputCurrentLimit1.%X1 := #statFrame.%X10;
                                   #statOutputCurrentLimit1.%X0 := #statFrame.%X11;

                                   //current limit of output 2 (0% to 100% of nominal value)
                                   #statOutputCurrentLimit2.%X3 := #statFrame.%X12;
                                   #statOutputCurrentLimit2.%X2 := #statFrame.%X13;
                                   #statOutputCurrentLimit2.%X1 := #statFrame.%X14;
                                   #statOutputCurrentLimit2.%X0 := #statFrame.%X15;

                                   //current limit of output 3 (0% to 100% of nominal value)
                                   #statOutputCurrentLimit3.%X3 := #statFrame.%X16;
                                   #statOutputCurrentLimit3.%X2 := #statFrame.%X17;
                                   #statOutputCurrentLimit3.%X1 := #statFrame.%X18;
                                   #statOutputCurrentLimit3.%X0 := #statFrame.%X19;

                                   //current limit of output 4 (0% to 100% of nominal value)
                                   #statOutputCurrentLimit4.%X3 := #statFrame.%X20;
                                   #statOutputCurrentLimit4.%X2 := #statFrame.%X21;
                                   #statOutputCurrentLimit4.%X1 := #statFrame.%X22;
                                   #statOutputCurrentLimit4.%X0 := #statFrame.%X23;

                               END_IF;

                               // state DIP switch
                               #statStateDipSwitchTD.%X1 := #statFrame.%X26;
                               #statHMI.stateDipSwitchTD1 := #statFrame.%X26;
                               #statStateDipSwitchTD.%X0 := #statFrame.%X27;
                               #statHMI.stateDipSwitchTD2 := #statFrame.%X27;


                               //0:= load dependent startup
                               //1:= startup time lag 25ms
                               //2:= startup time lag 250ms
                               //3:= startup time lag 500ms
                               #statHMI.startup := BYTE_TO_INT(#statStateDipSwitchTD);

                               //nominal output current
                               #statNominalOutputCurrent.%X1 := #statFrame.%X28;
                               #statNominalOutputCurrent.%X0 := #statFrame.%X29;


                               IF BYTE_TO_INT(#statNominalOutputCurrent) = #CONST_NOMINAL_VALUE_DETECT0
                               THEN
                                   #statHMI.nominalOutputCurrent := #CONST_NOMINAL_CURRENT3;
                               ELSIF BYTE_TO_INT(#statNominalOutputCurrent) = #CONST_NOMINAL_VALUE_DETECT1
                               THEN
                                   #statHMI.nominalOutputCurrent := #CONST_NOMINAL_CURRENT5;
                               ELSIF BYTE_TO_INT(#statNominalOutputCurrent) = #CONST_NOMINAL_VALUE_DETECT2
                               THEN
                                   #statHMI.nominalOutputCurrent := #CONST_NOMINAL_CURRENT10;
                               ELSE
                                   //default value
                                   #statHMI.nominalOutputCurrent := #CONST_NOMINAL_CURRENT3;

                               END_IF;

                               //number of outputs
                               IF #statFrame.%X30 = TRUE
                               THEN
                                   #statHMI.outputNumber := #CONST_OUTPUT_NUMBER_8;
                               ELSE
                                   #statHMI.outputNumber := #CONST_OUTPUT_NUMBER_4;
                               END_IF;

                               #statPower := #statHMI.nominalOutputCurrent * #CONST_NOMINAL_VOLTAGE * #statHMI.outputNumber;

                               // article number pos 7
                               IF #statPower > #CONST_POWER_0
                                   AND #statPower <= #CONST_POWER_20
                               THEN
                                   #statArticleNumber[7] := '0';
                               ELSIF #statPower > #CONST_POWER_20
                                   AND #statPower <= #CONST_POWER_50
                               THEN
                                   #statArticleNumber[7] := '1';
                               ELSIF #statPower > #CONST_POWER_50
                                   AND #statPower <= #CONST_POWER_100
                               THEN
                                   #statArticleNumber[7] := '2';
                               ELSIF #statPower > #CONST_POWER_100
                                   AND #statPower <= #CONST_POWER_150
                               THEN
                                   #statArticleNumber[7] := '3';
                               ELSIF #statPower > #CONST_POWER_150
                                   AND #statPower <= #CONST_POWER_250
                               THEN
                                   #statArticleNumber[7] := '4';
                               ELSIF #statPower > #CONST_POWER_250
                                   AND #statPower <= #CONST_POWER_400
                               THEN
                                   #statArticleNumber[7] := '5';
                               ELSIF #statPower > #CONST_POWER_400
                                   AND #statPower <= #CONST_POWER_600
                               THEN
                                   #statArticleNumber[7] := '6';
                               ELSIF #statPower > #CONST_POWER_600
                                   AND #statPower <= #CONST_POWER_1000
                               THEN
                                   #statArticleNumber[7] := '7';
                               ELSIF #statPower > #CONST_POWER_1000
                               THEN
                                   #statArticleNumber[7] := '8';
                               ELSE
                                   //default value
                                   #statArticleNumber[7] := '3';
                               END_IF;


                               IF #statGetFrame.frame21 = TRUE
                               THEN
                                   #statGetFrame.frame21 := false;

                                   #statHMI.outputCurrent1 := (BYTE_TO_INT(#statOutputCurrent1) * #statHMI.nominalOutputCurrent) / #CONST_CONVERT_CURRENT;
                                   #statHMI.outputCurrent2 := (BYTE_TO_INT(#statOutputCurrent2) * #statHMI.nominalOutputCurrent) / #CONST_CONVERT_CURRENT;
                                   #statHMI.outputCurrent3 := (BYTE_TO_INT(#statOutputCurrent3) * #statHMI.nominalOutputCurrent) / #CONST_CONVERT_CURRENT;
                                   #statHMI.outputCurrent4 := (BYTE_TO_INT(#statOutputCurrent4) * #statHMI.nominalOutputCurrent) / #CONST_CONVERT_CURRENT;

                               END_IF;

                               IF #statGetFrame.frame22 = true
                               THEN
                                   #statGetFrame.frame22 := false;

                                   IF #statCntReason > 10
                                   THEN
                                       #statCntReason := 0;
                                   END_IF;

                                   IF #statCntCurrentLimit > 10
                                   THEN
                                       #statCntCurrentLimit := 0;
                                   END_IF;

                                   //current limit or reason for switch off output 1
                                   IF #statHMI.stateOutput1 = #CONST_STATE_OUT_AUTO_SWITCHED_OFF OR
                                       #statHMI.stateOutput1 = #CONST_STATE_OUT_RESET_POSSIBLE
                                   THEN
                                       #statHMI.reasonOutputSwitchedOff1 := BYTE_TO_INT(#statOutputCurrentLimit1);
                                       #statCntReason := #statCntReason + 1;

                                   ELSE
                                       #statHMI.outputCurrentLimit1 := (BYTE_TO_INT(#statOutputCurrentLimit1) * #statHMI.nominalOutputCurrent) / #CONST_CONVERT_CURRENT;
                                       #statCntCurrentLimit := #statCntCurrentLimit + 1;
                                   END_IF;

                                   //current limit or reason for switch off output 2
                                   IF #statHMI.stateOutput2 = #CONST_STATE_OUT_AUTO_SWITCHED_OFF OR
                                       #statHMI.stateOutput2 = #CONST_STATE_OUT_RESET_POSSIBLE
                                   THEN
                                       #statHMI.reasonOutputSwitchedOff2 := BYTE_TO_INT(#statOutputCurrentLimit2);
                                   ELSE
                                       #statHMI.outputCurrentLimit2 := (BYTE_TO_INT(#statOutputCurrentLimit2) * #statHMI.nominalOutputCurrent) / #CONST_CONVERT_CURRENT;
                                   END_IF;

                                   //current limit or reason for switch off output 3
                                   IF #statHMI.stateOutput3 = #CONST_STATE_OUT_AUTO_SWITCHED_OFF OR
                                       #statHMI.stateOutput3 = #CONST_STATE_OUT_RESET_POSSIBLE
                                   THEN
                                       #statHMI.reasonOutputSwitchedOff3 := BYTE_TO_INT(#statOutputCurrentLimit3);
                                   ELSE
                                       #statHMI.outputCurrentLimit3 := (BYTE_TO_INT(#statOutputCurrentLimit3) * #statHMI.nominalOutputCurrent) / #CONST_CONVERT_CURRENT;
                                   END_IF;

                                   //current limit or reason for switch off output 4
                                   IF #statHMI.stateOutput4 = #CONST_STATE_OUT_AUTO_SWITCHED_OFF OR
                                       #statHMI.stateOutput4 = #CONST_STATE_OUT_RESET_POSSIBLE
                                   THEN
                                       #statHMI.reasonOutputSwitchedOff4 := BYTE_TO_INT(#statOutputCurrentLimit4);
                                   ELSE
                                       #statHMI.outputCurrentLimit4 := (BYTE_TO_INT(#statOutputCurrentLimit4) * #statHMI.nominalOutputCurrent) / #CONST_CONVERT_CURRENT;
                                   END_IF;

                               END_IF;

                           ELSIF BYTE_TO_INT(#statFrameID) = #CONST_FRAME_ID3
                           THEN

                               //measurements channel 5 to 8
                               #statGetFrame.frame3 := true;

                               #statMeasurementsChannels.%X1 := #statFrame.%X6;
                               #statMeasurementsChannels.%X0 := #statFrame.%X7;

                               IF BYTE_TO_INT(#statMeasurementsChannels) = #CONST_MEASUREMENT_CURRENT
                               THEN
                                   //measurement out current (channel 5 to 8)
                                   #statGetFrame.frame31 := true;

                                   //current output 5 (0% to 150% of nominal value)
                                   #statOutputCurrent5.%X3 := #statFrame.%X8;
                                   #statOutputCurrent5.%X2 := #statFrame.%X9;
                                   #statOutputCurrent5.%X1 := #statFrame.%X10;
                                   #statOutputCurrent5.%X0 := #statFrame.%X11;

                                   //current output 6 (0% to 150% of nominal value)
                                   #statOutputCurrent6.%X3 := #statFrame.%X12;
                                   #statOutputCurrent6.%X2 := #statFrame.%X13;
                                   #statOutputCurrent6.%X1 := #statFrame.%X14;
                                   #statOutputCurrent6.%X0 := #statFrame.%X15;

                                   //current output 7 (0% to 150% of nominal value)
                                   #statOutputCurrent7.%X3 := #statFrame.%X16;
                                   #statOutputCurrent7.%X2 := #statFrame.%X17;
                                   #statOutputCurrent7.%X1 := #statFrame.%X18;
                                   #statOutputCurrent7.%X0 := #statFrame.%X19;

                                   //current output 8 (0% to 150% of nominal value)
                                   #statOutputCurrent8.%X3 := #statFrame.%X20;
                                   #statOutputCurrent8.%X2 := #statFrame.%X21;
                                   #statOutputCurrent8.%X1 := #statFrame.%X22;
                                   #statOutputCurrent8.%X0 := #statFrame.%X23;

                               ELSIF BYTE_TO_INT(#statMeasurementsChannels) = #CONST_MEASUREMENT_CURRENT_LIMIT
                               THEN
                                   //output current limit on potentiometer (channel 5 to 8)
                                   #statGetFrame.frame32 := true;

                                   //current limit of output 5 (0% to 100% of nominal value)
                                   #statOutputCurrentLimit5.%X3 := #statFrame.%X8;
                                   #statOutputCurrentLimit5.%X2 := #statFrame.%X9;
                                   #statOutputCurrentLimit5.%X1 := #statFrame.%X10;
                                   #statOutputCurrentLimit5.%X0 := #statFrame.%X11;

                                   //current limit of output 6 (0% to 100% of nominal value)
                                   #statOutputCurrentLimit6.%X3 := #statFrame.%X12;
                                   #statOutputCurrentLimit6.%X2 := #statFrame.%X13;
                                   #statOutputCurrentLimit6.%X1 := #statFrame.%X14;
                                   #statOutputCurrentLimit6.%X0 := #statFrame.%X15;

                                   //current limit of output 7 (0% to 100% of nominal value)
                                   #statOutputCurrentLimit7.%X3 := #statFrame.%X16;
                                   #statOutputCurrentLimit7.%X2 := #statFrame.%X17;
                                   #statOutputCurrentLimit7.%X1 := #statFrame.%X18;
                                   #statOutputCurrentLimit7.%X0 := #statFrame.%X19;

                                   //current limit of output 8 (0% to 100% of nominal value)
                                   #statOutputCurrentLimit8.%X3 := #statFrame.%X20;
                                   #statOutputCurrentLimit8.%X2 := #statFrame.%X21;
                                   #statOutputCurrentLimit8.%X1 := #statFrame.%X22;
                                   #statOutputCurrentLimit8.%X0 := #statFrame.%X23;

                               END_IF;

                               // state DIP switch
                               #statStateDipSwitchTD.%X1 := #statFrame.%X26;
                               #statHMI.stateDipSwitchTD1 := #statFrame.%X26;
                               #statStateDipSwitchTD.%X0 := #statFrame.%X27;
                               #statHMI.stateDipSwitchTD2 := #statFrame.%X27;

                               //0:= load dependent startup
                               //1:= startup time lag 25ms
                               //2:= startup time lag 250ms
                               //3:= startup time lag 500ms
                               #statHMI.startup := BYTE_TO_INT(#statStateDipSwitchTD);

                               //nominal output current
                               #statNominalOutputCurrent.%X1 := #statFrame.%X28;
                               #statNominalOutputCurrent.%X0 := #statFrame.%X29;

                               IF BYTE_TO_INT(#statNominalOutputCurrent) = #CONST_NOMINAL_VALUE_DETECT0
                               THEN
                                   #statHMI.nominalOutputCurrent := #CONST_NOMINAL_CURRENT3;
                               ELSIF BYTE_TO_INT(#statNominalOutputCurrent) = #CONST_NOMINAL_VALUE_DETECT1
                               THEN
                                   #statHMI.nominalOutputCurrent := #CONST_NOMINAL_CURRENT5;
                               ELSIF BYTE_TO_INT(#statNominalOutputCurrent) = #CONST_NOMINAL_VALUE_DETECT2
                               THEN
                                   ;
                                   #statHMI.nominalOutputCurrent := #CONST_NOMINAL_CURRENT10;
                               ELSE
                                   //default value
                                   #statHMI.nominalOutputCurrent := #CONST_NOMINAL_CURRENT3;
                               END_IF;

                               //number of outputs
                               IF #statFrame.%X30 = TRUE
                               THEN
                                   #statHMI.outputNumber := #CONST_OUTPUT_NUMBER_8;
                               ELSE
                                   #statHMI.outputNumber := #CONST_OUTPUT_NUMBER_4;
                               END_IF;

                               IF #statGetFrame.frame31 = TRUE
                               THEN
                                   #statGetFrame.frame31 := false;

                                   #statHMI.outputCurrent5 := (BYTE_TO_INT(#statOutputCurrent5) * #statHMI.nominalOutputCurrent) / #CONST_CONVERT_CURRENT;
                                   #statHMI.outputCurrent6 := (BYTE_TO_INT(#statOutputCurrent6) * #statHMI.nominalOutputCurrent) / #CONST_CONVERT_CURRENT;
                                   #statHMI.outputCurrent7 := (BYTE_TO_INT(#statOutputCurrent7) * #statHMI.nominalOutputCurrent) / #CONST_CONVERT_CURRENT;
                                   #statHMI.outputCurrent8 := (BYTE_TO_INT(#statOutputCurrent8) * #statHMI.nominalOutputCurrent) / #CONST_CONVERT_CURRENT;

                               END_IF;

                               IF #statGetFrame.frame32 = TRUE
                               THEN
                                   #statGetFrame.frame32 := false;

                                   //current limit or reason for switch off output 5
                                   IF #statHMI.stateOutput5 = #CONST_STATE_OUT_AUTO_SWITCHED_OFF OR
                                       #statHMI.stateOutput5 = #CONST_STATE_OUT_RESET_POSSIBLE
                                   THEN
                                       #statHMI.reasonOutputSwitchedOff5 := #statOutputCurrentLimit5;
                                   ELSE
                                       #statHMI.outputCurrentLimit5 := (BYTE_TO_INT(#statOutputCurrentLimit5) * #statHMI.nominalOutputCurrent) / #CONST_CONVERT_CURRENT;
                                   END_IF;

